// TIA Portal project "HEAT-1-CADIZ-V15" (V20) (continued)

DATA_BLOCK "SafetyRobotDb"   // DB3, F_DB
{ S7_Optimized_Access := 'TRUE' }
VERSION : 0.1
BEGIN
END_DATA_BLOCK

// folder: Eliminar

DATA_BLOCK "DB_Supervisor"   // DB9
{ S7_Optimized_Access := 'TRUE' }
VERSION : 0.1
   VAR
      Common : Struct
         plc_ok : Bool;
         supervisor_ok : Bool;
         system_ok : Bool;
         safety_ok : Bool;
         air_ok : Bool;
         insp_water_ok : Bool;
         tank_water_ok : Bool;
         robot_ok : Bool;
         step_plc : Int;
         step_supervisor : Int;
         error : Bool;
         reset_req : Bool;
      END_STRUCT;
      Identification : Struct   // pag 2
         carriage_id_req : Bool;   // Sup->PLC
         new_carriage_id : Bool;   // PLC->Sup
         id_req : Bool;   // Sup->PLC
         id_running : Bool;   // PLC->Sup
         id_ok : Bool;   // PLC->Sup
         teach_req : Bool;   // Sup->PLC
         system_ok : Bool;   // PLC->Sup (parte de id_ok)
         pa_check_req : Bool;   // Sup->PLC
         tcg_req : Bool;   // Sup->PLC
      END_STRUCT;
      Teaching : Struct   // pag 3
         teach_ready : Bool;   // PLC->Sup
         teach_running : Bool;   // Sup->PLC
         teach_state : Bool;   // Sup->PLC
         jump_start_us : Bool;   // PLC->Sup
      END_STRUCT;
      StartUs : Struct   // pag 4
         start_us_ready : Bool;   // PLC->Sup
         start_us_running : Bool;   // Sup->PLC
         start_us_state : Bool;   // Sup->PLC
      END_STRUCT;
      PACheck : Struct   // pag 5
         pa_check_ready : Bool;   // PLC->Sup
         elem_running : Bool;   // Sup->PLC
         elem_state : Bool;   // Sup->PLC
         bal_running : Bool;   // Sup->PLC
         bal_state : Bool;   // Sup->PLC
      END_STRUCT;
      Gain : Struct
         gain_ready : Bool;
         gain_running : Bool;
         gain_state : Bool;
      END_STRUCT;
      TCG_Check : Struct
         tcg_ready : Bool;
         tcg_running : Bool;
         tcg_next_step : Bool;
         jump_acq_ref : Bool;
         jump_tcg_adj : Bool;
      END_STRUCT;
      TCG_Adjust : Struct
         tcg_ready : Bool;
         jump_ref_acq : Bool;
      END_STRUCT;
      RefScan_Acq : Struct
         scan_ref_ready : Bool;
         scan_ref_running : Bool;
      END_STRUCT;
      InspScan : Struct
         scan_insp_ready : Bool;
         scan_insp_running : Bool;
         scan_insp_state : Bool;
         jump_ref_insp : Bool;
      END_STRUCT;
      RefScan_Verif : Struct
         scan_ref_ready : Bool;
         scan_ref_running : Bool;
         jump_start : Bool;
      END_STRUCT;
      Marking : Struct
         mark_req : Bool;
         mark_running : Bool;
         mark_state : Bool;
         jump_start : Bool;
         point_coordinates : Struct
            x : Real;
            y : Real;
            z : Real;
            "a" : Real;
            "b" : Real;
            c : Real;
         END_STRUCT;
      END_STRUCT;
   END_VAR
BEGIN
END_DATA_BLOCK

// folder: 10. System

FUNCTION_BLOCK "SeqManager"   // FB20, LAD
{ S7_Optimized_Access := 'TRUE' }
VERSION : 0.1
   VAR_INPUT
      systemArmed : Bool;
      autoBusy : Bool;
      servBusy : Bool;
      teachingRunning : Bool;
      startUsRunning : Bool;
      modeRequest : UInt;
      modeReqSeq : UInt;
   END_VAR
   VAR_OUTPUT
      modeEffective : UInt;
      modeReady : Bool;
      enterService : Bool;
      enterAuto : Bool;
   END_VAR
   VAR
      lastSeq : UInt;
      safeAllOk : Bool;
      windowAuto : Bool;
      acceptSrv : Bool;
      acceptAuto : Bool;
   END_VAR
BEGIN

REGION Network 1 (SCL)
   #safeAllOk := #systemArmed;
   // Ventana AUTO: OR de todos los *_running (ver tablas por etapa en el PDF).  // nivel sostenido
   #windowAuto :=
   #teachingRunning OR #startUsRunning;

   #enterService := FALSE;
   #enterAuto := FALSE;
   #acceptSrv := FALSE;
   #acceptAuto := FALSE;
END_REGION

REGION Network 2 (SCL)
   // 1) Nueva petición por contador
   IF #modeReqSeq <> #lastSeq THEN
       #lastSeq := #modeReqSeq;

       CASE #modeRequest OF
           0:  // SERVICE
               IF #safeAllOk AND (NOT #autoBusy) AND (NOT #windowAuto) THEN
                   #acceptSrv := TRUE;
               END_IF;

           1:  // AUTO
               IF #safeAllOk AND (NOT #servBusy) THEN
                   #acceptAuto := TRUE;
               END_IF;

       END_CASE;
   END_IF;
END_REGION

REGION Network 3 (SCL)
   IF #acceptSrv THEN
       #modeEffective := 0;
       #enterService := TRUE;
   ELSIF #acceptAuto THEN
       #modeEffective := 1;
       #enterAuto := TRUE;
   END_IF;

   // 3) Ready hacia HMI
   IF #modeEffective = 0 THEN
       #modeReady := #safeAllOk AND (NOT #autoBusy);
   ELSE
       #modeReady := #safeAllOk AND (NOT #servBusy);
   END_IF;
END_REGION
END_FUNCTION_BLOCK

FUNCTION_BLOCK "KukaControlSeq"   // FB21, LAD
{ S7_Optimized_Access := 'TRUE' }
VERSION : 0.1
BEGIN

REGION Network 1: Envia posiciones a la aplicacion KukaControl
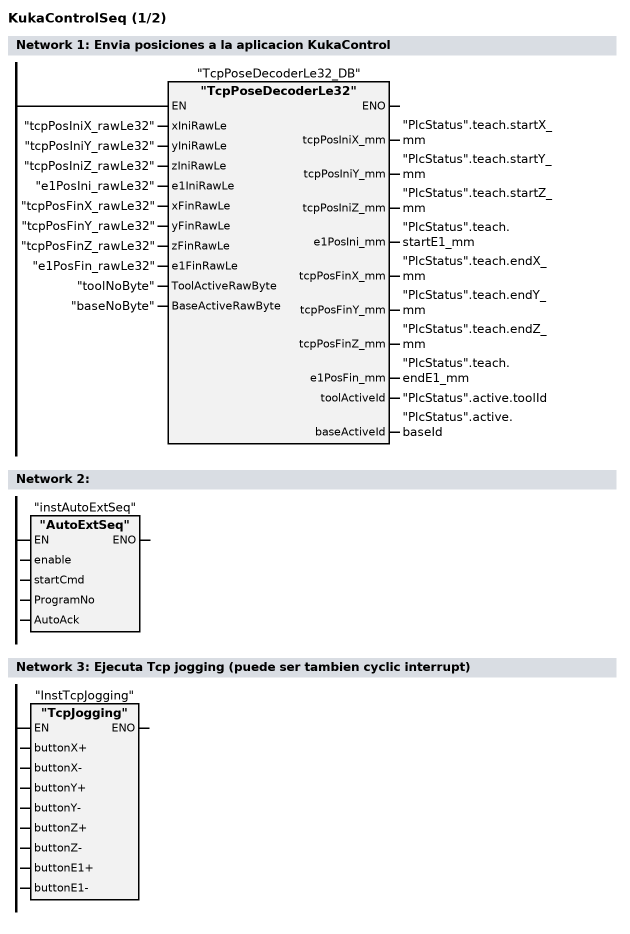
   RUNG wire#powerrail
      "TcpPoseDecoderLe32_DB"(xIniRawLe := "tcpPosIniX_rawLe32", yIniRawLe := "tcpPosIniY_rawLe32", zIniRawLe := "tcpPosIniZ_rawLe32", e1IniRawLe := "e1PosIni_rawLe32", xFinRawLe := "tcpPosFinX_rawLe32", yFinRawLe := "tcpPosFinY_rawLe32", zFinRawLe := "tcpPosFinZ_rawLe32", e1FinRawLe := "e1PosFin_rawLe32", ToolActiveRawByte := "toolNoByte", BaseActiveRawByte := "baseNoByte", tcpPosIniX_mm => "PlcStatus".teach.startX_mm, tcpPosIniY_mm => "PlcStatus".teach.startY_mm, tcpPosIniZ_mm => "PlcStatus".teach.startZ_mm, e1PosIni_mm => "PlcStatus".teach.startE1_mm, tcpPosFinX_mm => "PlcStatus".teach.endX_mm, tcpPosFinY_mm => "PlcStatus".teach.endY_mm, tcpPosFinZ_mm => "PlcStatus".teach.endZ_mm, e1PosFin_mm => "PlcStatus".teach.endE1_mm, toolActiveId => "PlcStatus".active.toolId, baseActiveId => "PlcStatus".active.baseId)
   END_RUNG
   // the same network as SCL:
   "TcpPoseDecoderLe32_DB"(xIniRawLe := "tcpPosIniX_rawLe32",   // "TcpPoseDecoderLe32"
                           yIniRawLe := "tcpPosIniY_rawLe32",
                           zIniRawLe := "tcpPosIniZ_rawLe32",
                           e1IniRawLe := "e1PosIni_rawLe32",
                           xFinRawLe := "tcpPosFinX_rawLe32",
                           yFinRawLe := "tcpPosFinY_rawLe32",
                           zFinRawLe := "tcpPosFinZ_rawLe32",
                           e1FinRawLe := "e1PosFin_rawLe32",
                           ToolActiveRawByte := "toolNoByte",
                           BaseActiveRawByte := "baseNoByte",
                           tcpPosIniX_mm => "PlcStatus".teach.startX_mm,
                           tcpPosIniY_mm => "PlcStatus".teach.startY_mm,
                           tcpPosIniZ_mm => "PlcStatus".teach.startZ_mm,
                           e1PosIni_mm => "PlcStatus".teach.startE1_mm,
                           tcpPosFinX_mm => "PlcStatus".teach.endX_mm,
                           tcpPosFinY_mm => "PlcStatus".teach.endY_mm,
                           tcpPosFinZ_mm => "PlcStatus".teach.endZ_mm,
                           e1PosFin_mm => "PlcStatus".teach.endE1_mm,
                           toolActiveId => "PlcStatus".active.toolId,
                           baseActiveId => "PlcStatus".active.baseId);
END_REGION

REGION Network 2
   RUNG wire#powerrail
      "instAutoExtSeq"(enable :=, startCmd :=, ProgramNo :=, AutoAck :=)
   END_RUNG
   // the same network as SCL:
   "instAutoExtSeq"();   // "AutoExtSeq"
END_REGION

REGION Network 3: Ejecuta Tcp jogging (puede ser tambien cyclic interrupt)
   RUNG wire#powerrail
      "InstTcpJogging"("buttonX+" :=, "buttonX-" :=, "buttonY+" :=, "buttonY-" :=, "buttonZ+" :=, "buttonZ-" :=, "buttonE1+" :=, "buttonE1-" :=)
   END_RUNG
   // the same network as SCL:
   "InstTcpJogging"();   // "TcpJogging"
END_REGION

REGION Network 4: Ejecuta TcpTarget
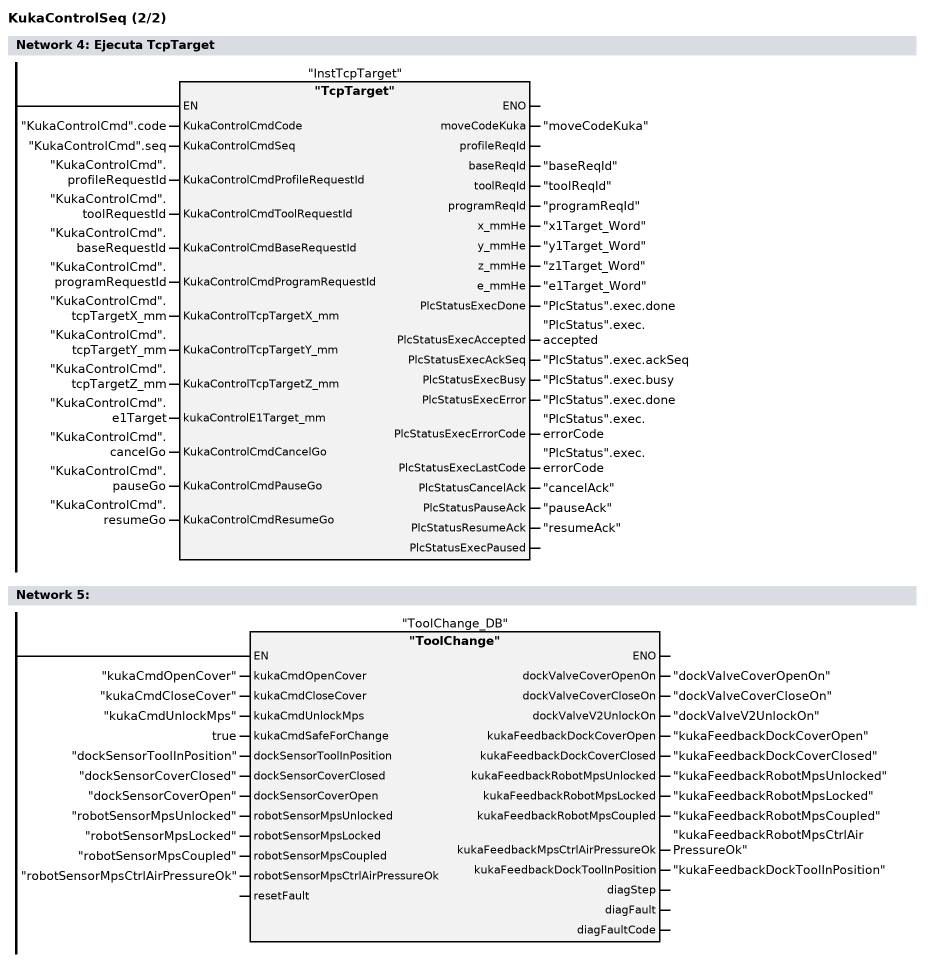
   RUNG wire#powerrail
      "InstTcpTarget"(KukaControlCmdCode := "KukaControlCmd".code, KukaControlCmdSeq := "KukaControlCmd".seq, KukaControlCmdProfileRequestId := "KukaControlCmd".profileRequestId, KukaControlCmdToolRequestId := "KukaControlCmd".toolRequestId, KukaControlCmdBaseRequestId := "KukaControlCmd".baseRequestId, KukaControlCmdProgramRequestId := "KukaControlCmd".programRequestId, KukaControlTcpTargetX_mm := "KukaControlCmd".tcpTargetX_mm, KukaControlTcpTargetY_mm := "KukaControlCmd".tcpTargetY_mm, KukaControlTcpTargetZ_mm := "KukaControlCmd".tcpTargetZ_mm, kukaControlE1Target_mm := "KukaControlCmd".e1Target, KukaControlCmdCancelGo := "KukaControlCmd".cancelGo, KukaControlCmdPauseGo := "KukaControlCmd".pauseGo, KukaControlCmdResumeGo := "KukaControlCmd".resumeGo, moveCodeKuka => "moveCodeKuka", profileReqId =>, baseReqId => "baseReqId", toolReqId => "toolReqId", programReqId => "programReqId", x_mmHe => "x1Target_Word", y_mmHe => "y1Target_Word", z_mmHe => "z1Target_Word", e_mmHe => "e1Target_Word", PlcStatusExecDone => "PlcStatus".exec.done, PlcStatusExecAccepted => "PlcStatus".exec.accepted, PlcStatusExecAckSeq => "PlcStatus".exec.ackSeq, PlcStatusExecBusy => "PlcStatus".exec.busy, PlcStatusExecError => "PlcStatus".exec.done, PlcStatusExecErrorCode => "PlcStatus".exec.errorCode, PlcStatusExecLastCode => "PlcStatus".exec.errorCode, PlcStatusCancelAck => "cancelAck", PlcStatusPauseAck => "pauseAck", PlcStatusResumeAck => "resumeAck", PlcStatusExecPaused =>)
   END_RUNG
   // the same network as SCL:
   "InstTcpTarget"(KukaControlCmdCode := "KukaControlCmd".code,   // "TcpTarget"
                   KukaControlCmdSeq := "KukaControlCmd".seq,
                   KukaControlCmdProfileRequestId := "KukaControlCmd".profileRequestId,
                   KukaControlCmdToolRequestId := "KukaControlCmd".toolRequestId,
                   KukaControlCmdBaseRequestId := "KukaControlCmd".baseRequestId,
                   KukaControlCmdProgramRequestId := "KukaControlCmd".programRequestId,
                   KukaControlTcpTargetX_mm := "KukaControlCmd".tcpTargetX_mm,
                   KukaControlTcpTargetY_mm := "KukaControlCmd".tcpTargetY_mm,
                   KukaControlTcpTargetZ_mm := "KukaControlCmd".tcpTargetZ_mm,
                   kukaControlE1Target_mm := "KukaControlCmd".e1Target,
                   KukaControlCmdCancelGo := "KukaControlCmd".cancelGo,
                   KukaControlCmdPauseGo := "KukaControlCmd".pauseGo,
                   KukaControlCmdResumeGo := "KukaControlCmd".resumeGo,
                   moveCodeKuka => "moveCodeKuka",
                   baseReqId => "baseReqId",
                   toolReqId => "toolReqId",
                   programReqId => "programReqId",
                   x_mmHe => "x1Target_Word",
                   y_mmHe => "y1Target_Word",
                   z_mmHe => "z1Target_Word",
                   e_mmHe => "e1Target_Word",
                   PlcStatusExecDone => "PlcStatus".exec.done,
                   PlcStatusExecAccepted => "PlcStatus".exec.accepted,
                   PlcStatusExecAckSeq => "PlcStatus".exec.ackSeq,
                   PlcStatusExecBusy => "PlcStatus".exec.busy,
                   PlcStatusExecError => "PlcStatus".exec.done,
                   PlcStatusExecErrorCode => "PlcStatus".exec.errorCode,
                   PlcStatusExecLastCode => "PlcStatus".exec.errorCode,
                   PlcStatusCancelAck => "cancelAck",
                   PlcStatusPauseAck => "pauseAck",
                   PlcStatusResumeAck => "resumeAck");
END_REGION

REGION Network 5
   RUNG wire#powerrail
      "ToolChange_DB"(kukaCmdOpenCover := "kukaCmdOpenCover", kukaCmdCloseCover := "kukaCmdCloseCover", kukaCmdUnlockMps := "kukaCmdUnlockMps", kukaCmdSafeForChange := true, dockSensorToolInPosition := "dockSensorToolInPosition", dockSensorCoverClosed := "dockSensorCoverClosed", dockSensorCoverOpen := "dockSensorCoverOpen", robotSensorMpsUnlocked := "robotSensorMpsUnlocked", robotSensorMpsLocked := "robotSensorMpsLocked", robotSensorMpsCoupled := "robotSensorMpsCoupled", robotSensorMpsCtrlAirPressureOk := "robotSensorMpsCtrlAirPressureOk", resetFault :=, dockValveCoverOpenOn => "dockValveCoverOpenOn", dockValveCoverCloseOn => "dockValveCoverCloseOn", dockValveV2UnlockOn => "dockValveV2UnlockOn", kukaFeedbackDockCoverOpen => "kukaFeedbackDockCoverOpen", kukaFeedbackDockCoverClosed => "kukaFeedbackDockCoverClosed", kukaFeedbackRobotMpsUnlocked => "kukaFeedbackRobotMpsUnlocked", kukaFeedbackRobotMpsLocked => "kukaFeedbackRobotMpsLocked", kukaFeedbackRobotMpsCoupled => "kukaFeedbackRobotMpsCoupled", kukaFeedbackMpsCtrlAirPressureOk => "kukaFeedbackRobotMpsCtrlAirPressureOk", kukaFeedbackDockToolInPosition => "kukaFeedbackDockToolInPosition", diagStep =>, diagFault =>, diagFaultCode =>)
   END_RUNG
   // the same network as SCL:
   "ToolChange_DB"(kukaCmdOpenCover := "kukaCmdOpenCover",   // "ToolChange"
                   kukaCmdCloseCover := "kukaCmdCloseCover",
                   kukaCmdUnlockMps := "kukaCmdUnlockMps",
                   kukaCmdSafeForChange := true,
                   dockSensorToolInPosition := "dockSensorToolInPosition",
                   dockSensorCoverClosed := "dockSensorCoverClosed",
                   dockSensorCoverOpen := "dockSensorCoverOpen",
                   robotSensorMpsUnlocked := "robotSensorMpsUnlocked",
                   robotSensorMpsLocked := "robotSensorMpsLocked",
                   robotSensorMpsCoupled := "robotSensorMpsCoupled",
                   robotSensorMpsCtrlAirPressureOk := "robotSensorMpsCtrlAirPressureOk",
                   dockValveCoverOpenOn => "dockValveCoverOpenOn",
                   dockValveCoverCloseOn => "dockValveCoverCloseOn",
                   dockValveV2UnlockOn => "dockValveV2UnlockOn",
                   kukaFeedbackDockCoverOpen => "kukaFeedbackDockCoverOpen",
                   kukaFeedbackDockCoverClosed => "kukaFeedbackDockCoverClosed",
                   kukaFeedbackRobotMpsUnlocked => "kukaFeedbackRobotMpsUnlocked",
                   kukaFeedbackRobotMpsLocked => "kukaFeedbackRobotMpsLocked",
                   kukaFeedbackRobotMpsCoupled => "kukaFeedbackRobotMpsCoupled",
                   kukaFeedbackMpsCtrlAirPressureOk => "kukaFeedbackRobotMpsCtrlAirPressureOk",
                   kukaFeedbackDockToolInPosition => "kukaFeedbackDockToolInPosition");
END_REGION
END_FUNCTION_BLOCK

FUNCTION_BLOCK "SupervisorSeq"   // FB22, LAD
{ S7_Optimized_Access := 'TRUE' }
VERSION : 0.1
   VAR
      firstScan : Bool;
      enteredStep : Bool;
      prev_step_plc : Int;
      prev_step_supervisor : Int;
      phase : Int;
      tcg_pos_index : Int;
      tcg_gate : Bool;
      cStep_IDENT : Int;
      cSTEP_TEACH : Int;
      cSTEP_STARTUS : Int;
      cSTEP_PA_CHECK : Int;
      cSTEP_GAIN : Int;
      cSTEP_TCG_CHECK : Int;
      cSTEP_TCG_ADJ : Int;
      cSTEP_REF_ACQ : Int;
      cSTEP_INSP : Int;
      cSTEP_REF_VERIF : Int;
      cSTEP_MARKING : Int;
   END_VAR
BEGIN

REGION Network 1 (SCL)
   IF #firstScan THEN
       "PlcStatus".Supervisor.global.plcOk := TRUE;


       "DB_Supervisor".Common.plc_ok := TRUE;
       "DB_Supervisor".Common.step_plc := #cStep_IDENT;
       #firstScan := FALSE;
   END_IF;

   "DB_Supervisor".Common.plc_ok := TRUE;


   // ---- State machine ----

   CASE "SupervisorCmd".global.stepSupervisor OF
           // 1) Identification (p.2)
       1:

           "DB_Supervisor".Identification.new_carriage_id :=
           "DB_Supervisor".Identification.carriage_id_req;

           CASE #phase OF
               0:
                   IF "DB_Supervisor".Identification.id_req THEN
                       "DB_Supervisor".Identification.id_running := TRUE;
                       "DB_Supervisor".Identification.id_ok :=
                       "DB_Supervisor".Common.safety_ok
                       AND "DB_Supervisor".Common.air_ok
                       AND "DB_Supervisor".Common.insp_water_ok
                       AND "DB_Supervisor".Common.tank_water_ok
                       AND "DB_Supervisor".Common.robot_ok
                       AND "DB_Supervisor".Common.supervisor_ok
                       AND "DB_Supervisor".Identification.system_ok;
                       #phase := 1;
                   END_IF;
               1:
                   "DB_Supervisor".Identification.id_running := FALSE;
                   IF "DB_Supervisor".Identification.id_ok THEN
                       IF "DB_Supervisor".Identification.teach_req THEN
                           "DB_Supervisor".Common.step_plc := 2;
                       ELSE
                           "DB_Supervisor".Common.step_plc := 3;
                       END_IF;
                   END_IF;
           END_CASE;

           ;

           // 2) Teaching (p.3)
       2:

           CASE  #phase OF
               0:
                   "DB_Supervisor".Teaching.teach_ready := TRUE;
                   IF "DB_Supervisor".Teaching.teach_running THEN
                       "DB_Supervisor".Teaching.teach_ready := FALSE;
                       #phase := 1;
                   END_IF;
               1:
                   IF NOT "DB_Supervisor".Teaching.teach_running THEN
                       IF "DB_Supervisor".Teaching.teach_state THEN
                           "DB_Supervisor".Common.step_plc := 3;
                       END_IF;
                   END_IF;
           END_CASE;


           // 3) Start US (p.4)
           3:

           CASE #phase OF
               0:
                   "DB_Supervisor".StartUs.start_us_ready := TRUE;
                   IF "DB_Supervisor".StartUs.start_us_running THEN
                       "DB_Supervisor".StartUs.start_us_ready := FALSE;
                       #phase := 1;
                   END_IF;
               1:
                   IF NOT "DB_Supervisor".StartUs.start_us_running THEN
                       IF "DB_Supervisor".StartUs.start_us_state THEN
                           IF "DB_Supervisor".Identification.pa_check_req THEN
                               "DB_Supervisor".Common.step_plc := 4;
                           ELSE
                               "DB_Supervisor".Common.step_plc := 5;
                           END_IF;
                       END_IF;
                   END_IF;
           END_CASE;


           // 4) PA‑Check (p.5)
           4:

           CASE #phase OF
               0:
                   "DB_Supervisor".PACheck.pa_check_ready := TRUE;
                   IF "DB_Supervisor".PACheck.elem_running THEN
                       "DB_Supervisor".PACheck.pa_check_ready := FALSE;
                       #phase := 1;
                   END_IF;
               1:
                   IF NOT "DB_Supervisor".PACheck.elem_running THEN
                       IF "DB_Supervisor".PACheck.elem_state THEN
                           #phase := 2;
                       END_IF;
                   END_IF;
               2:
                   IF "DB_Supervisor".PACheck.bal_running THEN
                       #phase := 3;
                   END_IF;
               3:
                   IF NOT "DB_Supervisor".PACheck.bal_running THEN
                       IF "DB_Supervisor".PACheck.bal_state THEN
                           "DB_Supervisor".Common.step_plc := 5;
                       END_IF;
                   END_IF;
           END_CASE;


           // 5) Gain (p.6)
           5:

           CASE #phase OF
               0:
                   "DB_Supervisor".Gain.gain_ready := TRUE;
                   IF "DB_Supervisor".Gain.gain_running THEN
                       "DB_Supervisor".Gain.gain_ready := FALSE;
                       #phase := 1;
                   END_IF;
               1:
                   IF NOT "DB_Supervisor".Gain.gain_running THEN
                       IF "DB_Supervisor".Gain.gain_state THEN
                           IF "DB_Supervisor".Identification.tcg_req THEN
                               "DB_Supervisor".Common.step_plc := 6;
                           ELSE
                               "DB_Supervisor".Common.step_plc := 8;
                           END_IF;
                       END_IF;
                   END_IF;
           END_CASE;


           // 6) TCG Check (p.7)
           6:

           CASE #phase OF
               0:
                   "DB_Supervisor".TCG_Check.tcg_ready := TRUE;
                   #tcg_pos_index := 0;
                   IF "DB_Supervisor".TCG_Check.tcg_running THEN
                       "DB_Supervisor".TCG_Check.tcg_ready := FALSE;
                       #phase := 1;
                   END_IF;

               1: // gate a tcg_next_step
                   IF "DB_Supervisor".TCG_Check.tcg_next_step AND NOT #tcg_gate THEN
                       #tcg_gate := TRUE;
                       #tcg_pos_index := #tcg_pos_index + 1; // 1..3
                   END_IF;
                   IF NOT "DB_Supervisor".TCG_Check.tcg_next_step THEN
                       #tcg_gate := FALSE;
                   END_IF;

                   IF NOT "DB_Supervisor".TCG_Check.tcg_running THEN
                       #phase := 2;
                   END_IF;

               2:
                   IF #tcg_pos_index >= 3 THEN
                       IF "DB_Supervisor".TCG_Check.jump_acq_ref THEN
                           "DB_Supervisor".Common.step_plc := 8;
                       ELSIF "DB_Supervisor".TCG_Check.jump_tcg_adj THEN
                           "DB_Supervisor".Common.step_plc := 7;
                       END_IF;
                   END_IF;
           END_CASE;


           // 7) TCG Adjust (p.7)
           7:

           CASE #phase OF
               0:
                   "DB_Supervisor".TCG_Adjust.tcg_ready := TRUE;
                   #phase := 1;
               1:
                   IF "DB_Supervisor".TCG_Adjust.jump_ref_acq THEN
                       "DB_Supervisor".Common.step_plc := 8;
                   END_IF;
           END_CASE;


           // 8) RefScan – Acquisition (p.8)
           8:

           CASE #phase OF
               0:
                   "DB_Supervisor".RefScan_Acq.scan_ref_ready := TRUE;
                   IF "DB_Supervisor".RefScan_Acq.scan_ref_running THEN
                       "DB_Supervisor".RefScan_Acq.scan_ref_ready := FALSE;
                       #phase := 1;
                   END_IF;
               1:
                   IF NOT "DB_Supervisor".RefScan_Acq.scan_ref_running THEN
                       "DB_Supervisor".Common.step_plc := 9;
                   END_IF;
           END_CASE;


           // 9) Inspection Scan (p.9)
           9:

           CASE #phase OF
               0:
                   "DB_Supervisor".InspScan.scan_insp_ready := TRUE;
                   IF "DB_Supervisor".InspScan.scan_insp_running THEN
                       "DB_Supervisor".InspScan.scan_insp_ready := FALSE;
                       #phase := 1;
                   END_IF;
               1:
                   IF "DB_Supervisor".InspScan.jump_ref_insp THEN
                       "DB_Supervisor".Common.step_plc := 10;
                   END_IF;
           END_CASE;


           // 10) RefScan – Verification (p.10)
           10:

           CASE #phase OF
               0:
                   "DB_Supervisor".RefScan_Verif.scan_ref_ready := TRUE;
                   IF "DB_Supervisor".RefScan_Verif.scan_ref_running THEN
                       "DB_Supervisor".RefScan_Verif.scan_ref_ready := FALSE;
                       #phase := 1;
                   END_IF;
               1:
                   IF "DB_Supervisor".RefScan_Verif.jump_start THEN
                       "DB_Supervisor".Common.step_plc := 1;
                   END_IF;
           END_CASE;

           // 11) Marking / Pre‑evaluation (p.11)
           11:

           CASE #phase OF
               0:
                   IF "DB_Supervisor".Marking.mark_req THEN
                       "DB_Supervisor".Marking.mark_running := TRUE;
                       #phase := 1;
                   END_IF;
               1:
                   // Sustituir por DONE real:
                   IF TRUE THEN
                       "DB_Supervisor".Marking.mark_running := FALSE;
                       "DB_Supervisor".Marking.mark_state := TRUE;
                       #phase := 2;
                   END_IF;
               2:
                   IF "DB_Supervisor".Marking.jump_start THEN
                       "DB_Supervisor".Common.step_plc := 1;
                   END_IF;
           END_CASE;


       ELSE
           "DB_Supervisor".Common.step_plc := 1;
       END_CASE;
END_REGION
END_FUNCTION_BLOCK

ORGANIZATION_BLOCK "Main"   // OB1, LAD, ProgramCycle
TITLE = "Main Program Sweep (Cycle)"
{ S7_Optimized_Access := 'TRUE' }
VERSION : 0.1
   VAR_INPUT
      Initial_Call : Bool;   // Initial call of this OB
      Remanence : Bool;   // =True, if remanent data are available
   END_VAR
   VAR_TEMP
      evtEnterSrv : Bool;   // // Eventos de modo service jog
      evtEnterAuto : Bool;   // // Eventos de modo auto
      muxSelStb : Bool;
      muxStartStb : Bool;
      muxPgno : Byte;
      u : UDInt;
   END_VAR
BEGIN

REGION Network 1 (SCL): // ====================== READ (%I) ======================
   // // —— Enlaza estos símbolos a tus %I en el árbol de dispositivos ——
   //   // EStop_DI, SafeDoor_DI, AirPressure_DI, WaterInsp_DI, WaterTank_DI, RobotReady_DI, ...
END_REGION

REGION Network 2: // 1) Árbitro de modo: decide y emite
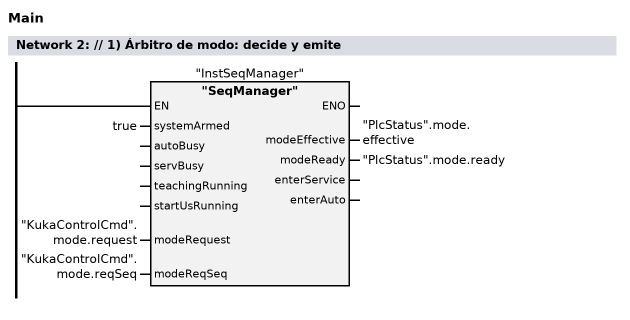
   RUNG wire#powerrail
      "InstSeqManager"(systemArmed := true, autoBusy :=, servBusy :=, teachingRunning :=, startUsRunning :=, modeRequest := "KukaControlCmd".mode.request, modeReqSeq := "KukaControlCmd".mode.reqSeq, modeEffective => "PlcStatus".mode.effective, modeReady => "PlcStatus".mode.ready, enterService =>, enterAuto =>)
   END_RUNG
   // the same network as SCL:
   "InstSeqManager"(systemArmed := true,   // "SeqManager"
                    modeRequest := "KukaControlCmd".mode.request,
                    modeReqSeq := "KukaControlCmd".mode.reqSeq,
                    modeEffective => "PlcStatus".mode.effective,
                    modeReady => "PlcStatus".mode.ready);
END_REGION

REGION Network 3 (SCL): // 2) Ejecuta o service o Auto
       IF "PlcStatus".mode.effective = 1 THEN
           // SUPERVISOR : Mode Effective = 1
           "InstSupervisorSeq"();
       ELSE
           // KUKACONTROL: Mode Effective = 0
           "InstKukaControlSeq"();
       END_IF;
END_REGION
END_ORGANIZATION_BLOCK

// folder: 10. System/Utilities

FUNCTION_BLOCK "ClockPulse"   // FB67, LAD
{ S7_Optimized_Access := 'TRUE' }
VERSION : 0.1
BEGIN
END_FUNCTION_BLOCK

// folder: 20. Robot Services/AutoExt

FUNCTION_BLOCK "AutoExtSeq"   // FB31, LAD
{ S7_Optimized_Access := 'TRUE' }
VERSION : 0.1
   VAR_INPUT
      enable : Bool;   // // habilita interfaz
      startCmd : Bool;   // // flanco de arranque
      ProgramNo : Byte;   // / nº CASE (1..255)
      AutoAck : Bool;   // // auto-confirmar STOPMESS
   END_VAR
   VAR
      rStart : R_TRIG;
      Static_1 : Bool;
      fReq : F_TRIG;
      pending : Bool;   // // hay pedido en curso
      running : Bool;   // // PRO_ACT latcheado
      pgnoLat : Byte;   // // PGNO latcheado
      tpStart : TP_TIME;
      tpAck : TP_TIME;
      rStop : R_TRIG;
   END_VAR
BEGIN

REGION Network 2 (SCL): // ---- detectar solicitud de arranque ----
END_REGION

REGION Network 3 (SCL): Paridad
END_REGION

REGION Network 4 (SCL): // ---- VALID solo mientras PGNO_REQ=1 y hay pedido ----
END_REGION

REGION Network 5 (SCL): // ---- cuando PGNO_REQ baja -> pulso de EXT_START ---
END_REGION

REGION Network 6 (SCL): // ---- auto-confirmar mensajes cuando aparezcan ----
END_REGION

REGION Network 7 (SCL): ---- seguimiento de ejecución y liberación de 'pending' ----
END_REGION
END_FUNCTION_BLOCK

// folder: 20. Robot Services/Mov Manual

FUNCTION_BLOCK "TcpJogging"   // FB5, LAD
{ S7_Optimized_Access := 'TRUE' }
VERSION : 0.1
   VAR_INPUT
      "buttonX+" : Bool;
      "buttonX-" : Bool;
      "buttonY+" : Bool;
      "buttonY-" : Bool;
      "buttonZ+" : Bool;
      "buttonZ-" : Bool;
      "buttonE1+" : Bool;
      "buttonE1-" : Bool;
   END_VAR
BEGIN

REGION Network 1 (SCL): Mapea los valores de los botones de WF
   IF "PlcStatus".mode.effective = 0 THEN

       "Tag_1" := TRUE;
       //MOV X,Y,Z
       //%Q630.0 = buttonX+
       //%Q630.1 = buttonX-
       //%Q630.2 = buttonY+
       //%Q630.3 = buttonY-
       //%Q630.4 = buttonZ+
       //%Q630.5 = buttonZ-
       //MOV A,B,C
       //%Q630.6 = buttonWF +A
       //%Q630.7 = buttonWF -A
       //%Q631.0 = buttonWF +B
       //%Q631.1 = buttonWF -B
       //%Q631.2 = buttonWF +C
       //%Q631.3 = buttonWF -C
       //Mov E1
       //%Q631.4 = buttonWF +E1
       //%Q631.5 = buttonWF -E1

   ELSE
       //%Q631.1 = buttonWF -B
       "Tag_1" := FALSE;
   END_IF;
END_REGION
END_FUNCTION_BLOCK

FUNCTION_BLOCK "TcpTarget"   // FB11, LAD
{ S7_Optimized_Access := 'TRUE' }
VERSION : 0.1
   VAR_INPUT
      KukaControlCmdCode : UInt;
      KukaControlCmdSeq : UInt;
      KukaControlCmdProfileRequestId : UInt;
      KukaControlCmdToolRequestId : UInt;
      KukaControlCmdBaseRequestId : UInt;
      KukaControlCmdProgramRequestId : UInt;
      KukaControlTcpTargetX_mm : LReal;
      KukaControlTcpTargetY_mm : LReal;
      KukaControlTcpTargetZ_mm : LReal;
      kukaControlE1Target_mm : LReal;
      KukaControlCmdCancelGo : Bool;
      KukaControlCmdPauseGo : Bool;
      KukaControlCmdResumeGo : Bool;
   END_VAR
   VAR_OUTPUT
      moveCodeKuka : Word;
      profileReqId : Word;
      baseReqId : Word;
      toolReqId : Word;
      programReqId : Word;
      x_mmHe : DWord;
      y_mmHe : DWord;
      z_mmHe : DWord;
      e_mmHe : DWord;
      PlcStatusExecDone : Bool;
      PlcStatusExecAccepted : Bool;
      PlcStatusExecAckSeq : UInt;
      PlcStatusExecBusy : Bool;
      PlcStatusExecError : Bool;
      PlcStatusExecErrorCode : DWord;
      PlcStatusExecLastCode : UInt;
      PlcStatusCancelAck : Bool;
      PlcStatusPauseAck : Bool;
      PlcStatusResumeAck : Bool;
      PlcStatusExecPaused : Bool;
   END_VAR
   VAR
      lastSeq : UInt;
      lastCode : UInt;
      state : Int;
      tmoMove : TON_TIME;
      rbDoneEdge : R_TRIG;
      _cancelInFlight : Bool := false;   // marca que el DONE que venga es por cancelación
      _isMotion : Bool;   // helper para saber si el code es de movimiento
   END_VAR
   VAR_TEMP
      x_dint : DInt;
      y_dint : DInt;
      z_dint : DInt;
      n_dint : DInt;
      code_int : UInt;
      tool_int : UInt;
   END_VAR
BEGIN

REGION Network 1 (SCL)
   // =================== Canal asíncrono ExecCtrl ====================
   // Handshake por nivel: <Go> de HMI -> PLC -> KRC, y cierre al recibir <Ack> del KRC.
   // Al cerrar, reflejamos el Ack hacia HMI y actualizamos PlcStatusExecPaused.

   // ---- CANCEL ----
   IF (#KukaControlCmdCancelGo <> #PlcStatusCancelAck) THEN
       "cancelGo" := #KukaControlCmdCancelGo;   // propaga al KRC
       #_cancelInFlight := TRUE;              // esperamos DONE por cancel
       // cerrar cuando el KRC confirme
       IF ("cancelAck" = "cancelGo") THEN
           #PlcStatusCancelAck := #KukaControlCmdCancelGo;  // cierra HMI
           #PlcStatusExecPaused := FALSE;                 // cancel limpia pausa (si la había)
       END_IF;
   END_IF;


   // ---- PAUSE ----
   IF (#KukaControlCmdPauseGo <> #PlcStatusPauseAck) THEN
       "pauseGo" := #KukaControlCmdPauseGo;     // propaga al KRC
       IF ("pauseAck" = "pauseGo") THEN
           #PlcStatusPauseAck := #KukaControlCmdPauseGo;    // cierra HMI
           #PlcStatusExecPaused := TRUE;                   // queda en pausa reanudable
       END_IF;
   END_IF;